(* Logix 5000 project; controller PLC_MCC1300_75F1 vendor 1 type 14 code 166 rev 32.11; software revision 32.04; part 50 of 83 *)
(* tags used below, declared in another part *)
   CM_ConveyorStackerToLine_JS1_Sync : CM_ConveyorStackerToLine;
   CONST_dDest_Cullet : DINT;
   CONST_dDest_Stk : DINT;
   CONST_rgdDestMask : DINT[32];   // Destination Mask
   Convoy_SL_DATA_NULL : UDT_Convoy_SL;
   GP_CheckIdPlatePresent : GP_CheckIdPlatePresent;
   GP_InvertCapxLite : GP_InvertCapxLite;
   GP_OB_InitializeMain : GP_OB_Initialize;
   GP_RampSpace : GP_RampSpace;
   Gp_SpaceConvUtilities_V1 : GP_SpaceConvUtilities_V1;
   M310B : MAC_Conveyor;
   M310B_ALM : MAC_Conveyor_ALM;
   M310B_Data : UDT_Convoy_SL;
   M310B_HMR : MAC_Conveyor_HMR;
   M310B_HMW : MAC_Conveyor_HMW;
   M310B_SpaceConv_Utilities : SpaceConv_Utilities;
   M310B_xPlateCullet : BOOL;
   M310Popup : MAC_Popup_ZC[2];
   M310Popup_SL_DATA : UDT_Convoy_SL;
   M311 : MAC_Conveyor;
   M311_Data : UDT_Convoy_SL;
   M311_SpaceConv_Utilities : SpaceConv_Utilities;
   M311_SpaceConvUtilities : SpaceConv_Utilities;
   M312 : MAC_Conveyor_Single;
   O : INT[128];
   TMP_d : DINT;
   TMP_dConveyorNumberForZoneCleaning : DINT;
   TMP_dDecelerationPositionEndConveyor : DINT;
   TMP_dHeadPosition : DINT;
   TMP_dOffsetLoadUnload_cmm : DINT;
   TMP_dPhEndPosition_cmm : DINT;
   TMP_dTailPosition : DINT;
   TMP_rgxId : DINT[10];
   TMP_SendToCullet : BOOL;
   TMP_xConveyorInvolvedInCleaning : BOOL;
   TMP_xConveyorOfStartCleaning : BOOL;
   TMP_xCulletPresent : BOOL;
   TMP_xEnableLoadUnload : BOOL;
   TMP_xEnableZoneCleaning : BOOL;
   TMP_xLiteThisDestPresent : BOOL;
   TMP_xReqUnpack : BOOL;
   xAlwaysOFF : BOOL;
   xAlwaysON : BOOL;
   Z401 : MAC_Zone;
   Z401_HMR : MAC_Zone_HMR;
   Z401_HMW : MAC_Zone_HMW;
(* MainProgram, continued *)

ROUTINE M310B_Logic   (* ladder *)
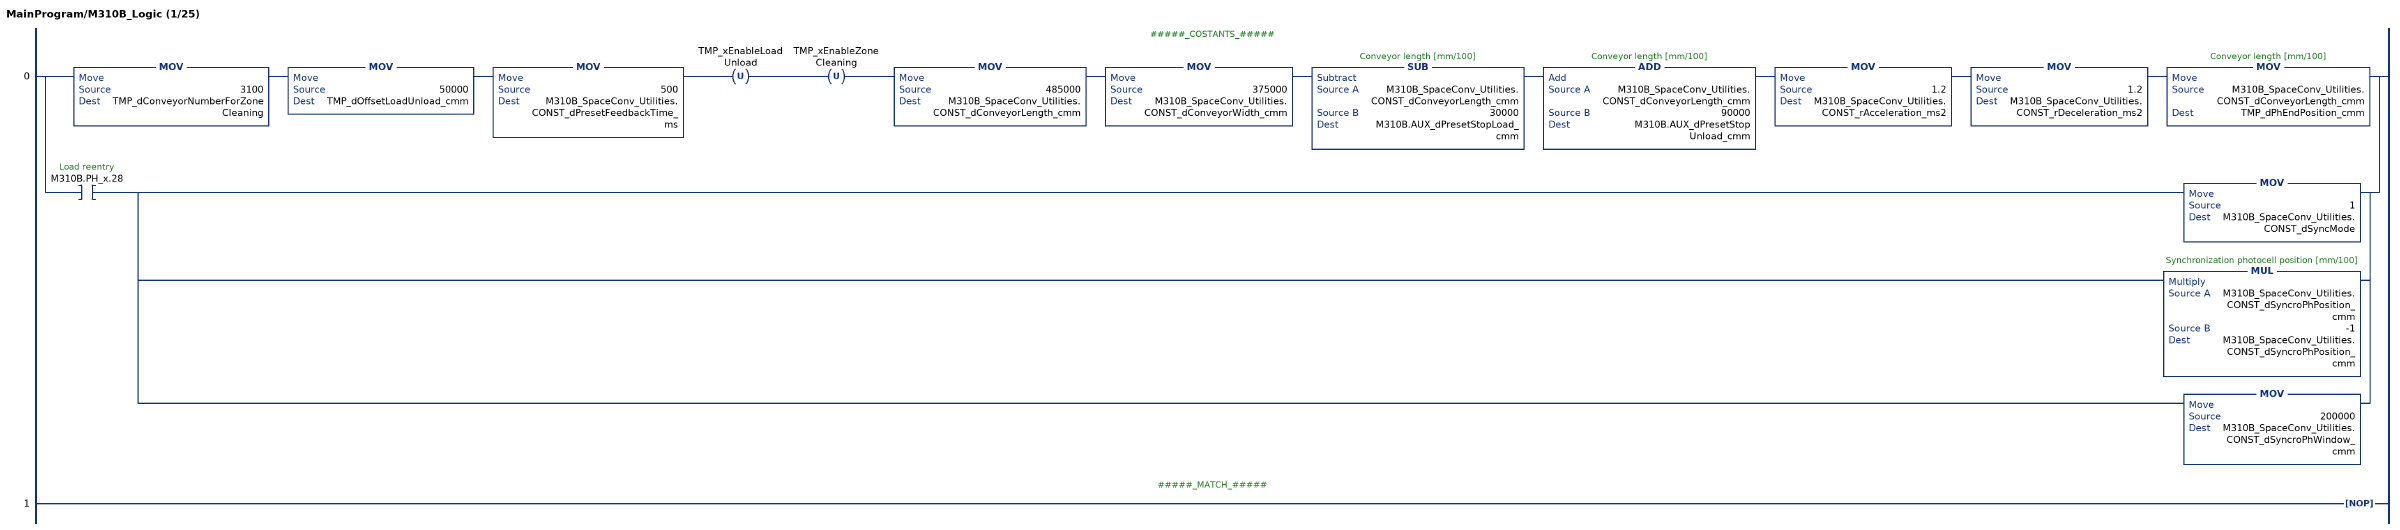
   // #####_COSTANTS_#####
   0: [MOV(3100,TMP_dConveyorNumberForZoneCleaning) MOV(50000,TMP_dOffsetLoadUnload_cmm) MOV(500,M310B_SpaceConv_Utilities.CONST_dPresetFeedbackTime_ms) OTU(TMP_xEnableLoadUnload) OTU(TMP_xEnableZoneCleaning) MOV(485000,M310B_SpaceConv_Utilities.CONST_dConveyorLength_cmm) MOV(375000,M310B_SpaceConv_Utilities.CONST_dConveyorWidth_cmm) SUB(M310B_SpaceConv_Utilities.CONST_dConveyorLength_cmm,30000,M310B.AUX_dPresetStopLoad_cmm) ADD(M310B_SpaceConv_Utilities.CONST_dConveyorLength_cmm,90000,M310B.AUX_dPresetStopUnload_cmm) MOV(1.2,M310B_SpaceConv_Utilities.CONST_rAcceleration_ms2) MOV(1.2,M310B_SpaceConv_Utilities.CONST_rDeceleration_ms2) MOV(M310B_SpaceConv_Utilities.CONST_dConveyorLength_cmm,TMP_dPhEndPosition_cmm) ,XIC(M310B.PH_x.28) [MOV(1,M310B_SpaceConv_Utilities.CONST_dSyncMode) ,MUL(M310B_SpaceConv_Utilities.CONST_dSyncroPhPosition_cmm,-1,M310B_SpaceConv_Utilities.CONST_dSyncroPhPosition_cmm) ,MOV(200000,M310B_SpaceConv_Utilities.CONST_dSyncroPhWindow_cmm) ] ];
   // #####_MATCH_#####
   1: NOP();
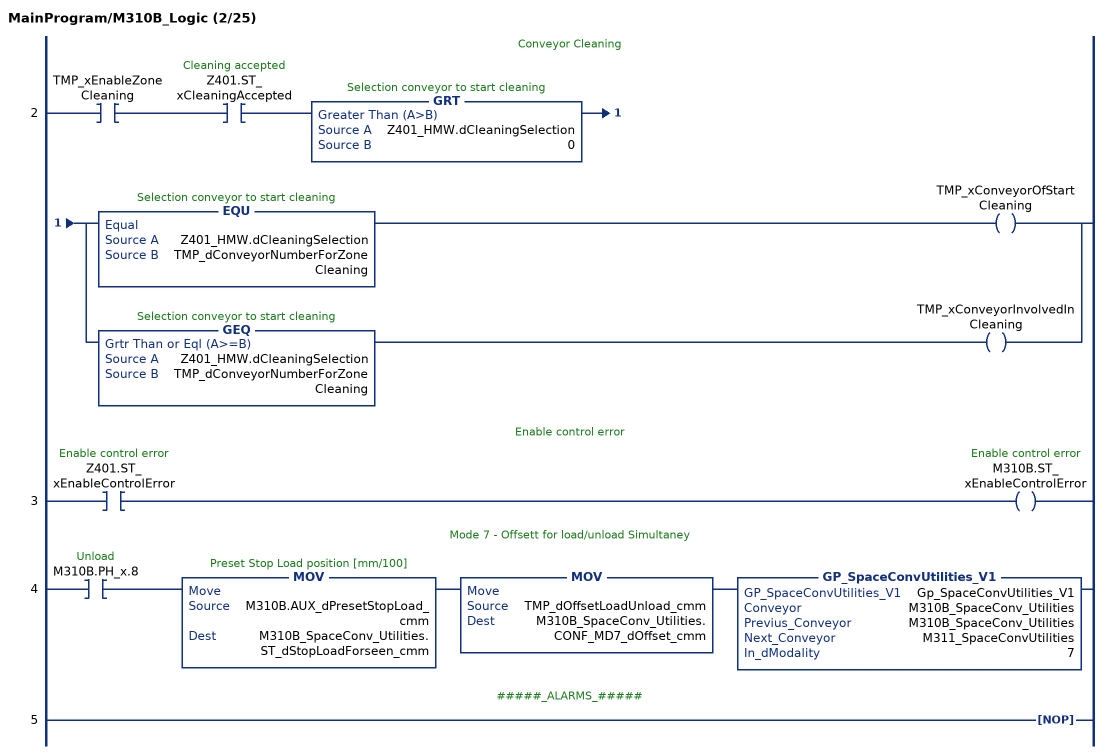
   // Conveyor Cleaning
   2: XIC(TMP_xEnableZoneCleaning)XIC(Z401.ST_xCleaningAccepted)GRT(Z401_HMW.dCleaningSelection,0)[EQU(Z401_HMW.dCleaningSelection,TMP_dConveyorNumberForZoneCleaning) OTE(TMP_xConveyorOfStartCleaning) ,GEQ(Z401_HMW.dCleaningSelection,TMP_dConveyorNumberForZoneCleaning) OTE(TMP_xConveyorInvolvedInCleaning) ];
   // Enable control error
   3: XIC(Z401.ST_xEnableControlError)OTE(M310B.ST_xEnableControlError);
   // Mode 7 - Offsett for load/unload Simultaney
   4: XIC(M310B.PH_x.8)MOV(M310B.AUX_dPresetStopLoad_cmm,M310B_SpaceConv_Utilities.ST_dStopLoadForseen_cmm)MOV(TMP_dOffsetLoadUnload_cmm,M310B_SpaceConv_Utilities.CONF_MD7_dOffset_cmm)GP_SpaceConvUtilities_V1(Gp_SpaceConvUtilities_V1,M310B_SpaceConv_Utilities,M310B_SpaceConv_Utilities,M311_SpaceConvUtilities,7);
   // #####_ALARMS_#####
   5: NOP();
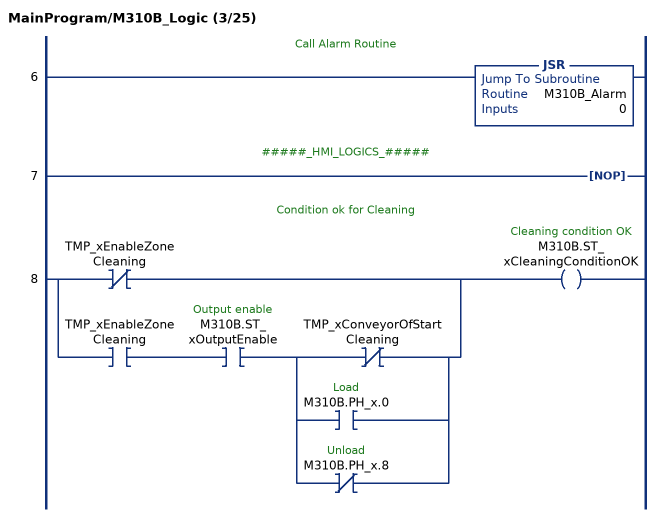
   // Call Alarm Routine
   6: JSR(M310B_Alarm,0);
   // #####_HMI_LOGICS_#####
   7: NOP();
   // Condition ok for Cleaning
   8: [XIO(TMP_xEnableZoneCleaning) ,XIC(TMP_xEnableZoneCleaning) XIC(M310B.ST_xOutputEnable) [XIO(TMP_xConveyorOfStartCleaning) ,XIC(M310B.PH_x.0) ,XIO(M310B.PH_x.8) ] ]OTE(M310B.ST_xCleaningConditionOK);
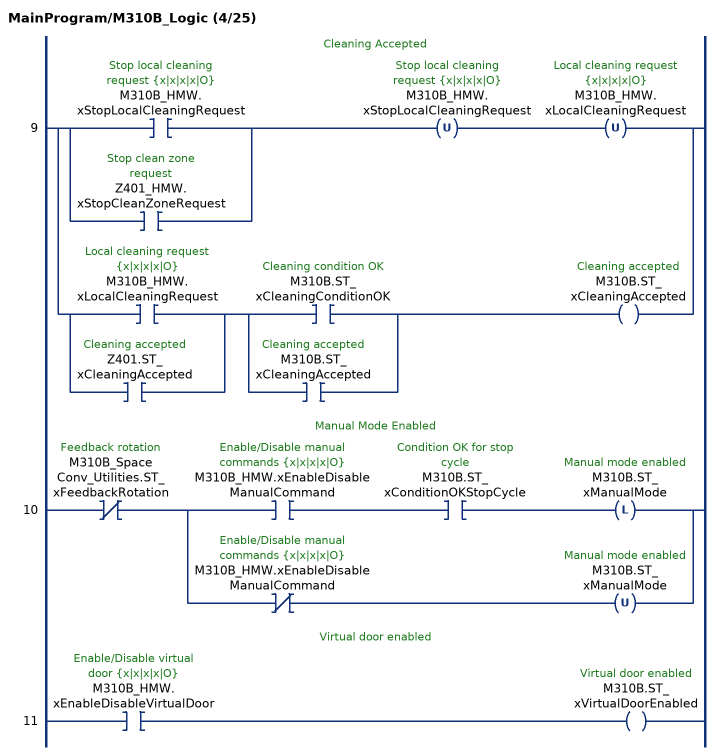
   // Cleaning Accepted
   9: [[XIC(M310B_HMW.xStopLocalCleaningRequest) ,XIC(Z401_HMW.xStopCleanZoneRequest) ] OTU(M310B_HMW.xStopLocalCleaningRequest) OTU(M310B_HMW.xLocalCleaningRequest) ,[XIC(M310B_HMW.xLocalCleaningRequest) ,XIC(Z401.ST_xCleaningAccepted) ] [XIC(M310B.ST_xCleaningConditionOK) ,XIC(M310B.ST_xCleaningAccepted) ] OTE(M310B.ST_xCleaningAccepted) ];
   // Manual Mode Enabled
   10: XIO(M310B_SpaceConv_Utilities.ST_xFeedbackRotation)[XIC(M310B_HMW.xEnableDisableManualCommand) XIC(M310B.ST_xConditionOKStopCycle) OTL(M310B.ST_xManualMode) ,XIO(M310B_HMW.xEnableDisableManualCommand) OTU(M310B.ST_xManualMode) ];
   // Virtual door enabled
   11: XIC(M310B_HMW.xEnableDisableVirtualDoor)OTE(M310B.ST_xVirtualDoorEnabled);
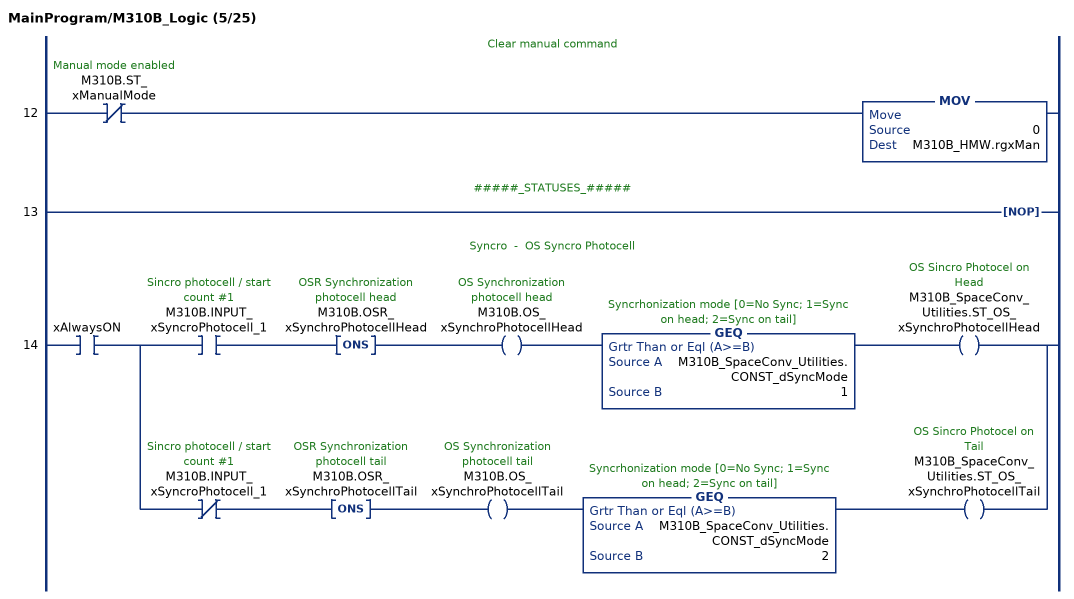
   // Clear manual command
   12: XIO(M310B.ST_xManualMode)MOV(0,M310B_HMW.rgxMan);
   // #####_STATUSES_#####
   13: NOP();
   // Syncro  -  OS Syncro Photocell
   14: XIC(xAlwaysON)[XIC(M310B.INPUT_xSyncroPhotocell_1) ONS(M310B.OSR_xSynchroPhotocellHead) OTE(M310B.OS_xSynchroPhotocellHead) GEQ(M310B_SpaceConv_Utilities.CONST_dSyncMode,1) OTE(M310B_SpaceConv_Utilities.ST_OS_xSynchroPhotocellHead) ,XIO(M310B.INPUT_xSyncroPhotocell_1) ONS(M310B.OSR_xSynchroPhotocellTail) OTE(M310B.OS_xSynchroPhotocellTail) GEQ(M310B_SpaceConv_Utilities.CONST_dSyncMode,2) OTE(M310B_SpaceConv_Utilities.ST_OS_xSynchroPhotocellTail) ];
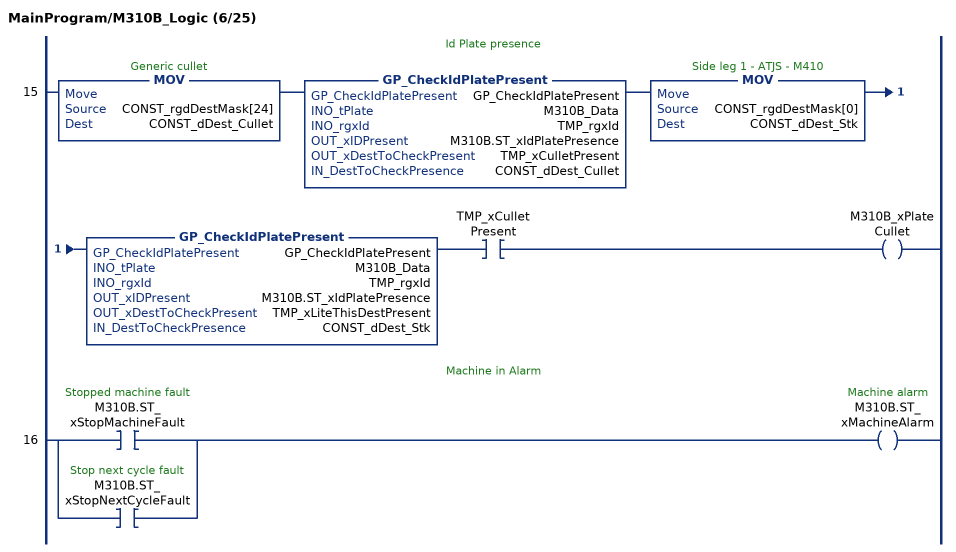
   // Id Plate presence
   15: MOV(CONST_rgdDestMask[24],CONST_dDest_Cullet)GP_CheckIdPlatePresent(GP_CheckIdPlatePresent,M310B_Data,TMP_rgxId,M310B.ST_xIdPlatePresence,TMP_xCulletPresent,CONST_dDest_Cullet)MOV(CONST_rgdDestMask[0],CONST_dDest_Stk)GP_CheckIdPlatePresent(GP_CheckIdPlatePresent,M310B_Data,TMP_rgxId,M310B.ST_xIdPlatePresence,TMP_xLiteThisDestPresent,CONST_dDest_Stk)XIC(TMP_xCulletPresent)OTE(M310B_xPlateCullet);
   // Machine in Alarm
   16: [XIC(M310B.ST_xStopMachineFault) ,XIC(M310B.ST_xStopNextCycleFault) ]OTE(M310B.ST_xMachineAlarm);
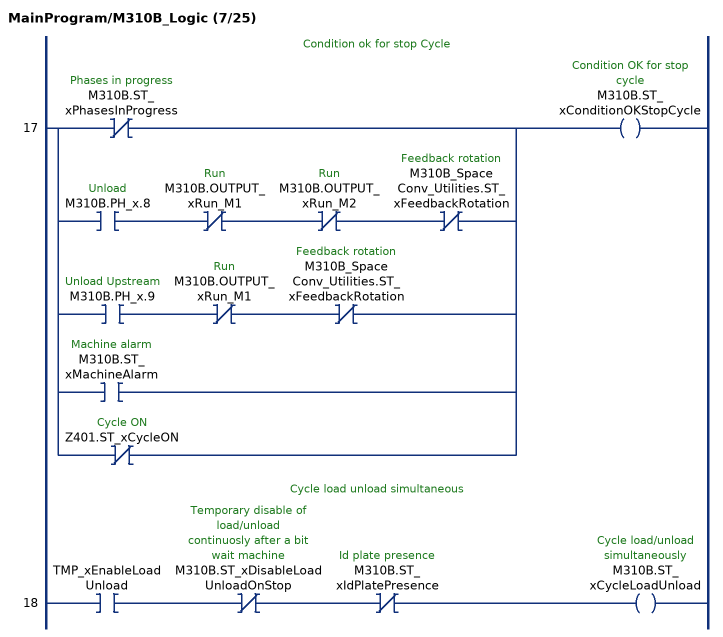
   // Condition ok for stop Cycle
   17: [XIO(M310B.ST_xPhasesInProgress) ,XIC(M310B.PH_x.8) XIO(M310B.OUTPUT_xRun_M1) XIO(M310B.OUTPUT_xRun_M2) XIO(M310B_SpaceConv_Utilities.ST_xFeedbackRotation) ,XIC(M310B.PH_x.9) XIO(M310B.OUTPUT_xRun_M1) XIO(M310B_SpaceConv_Utilities.ST_xFeedbackRotation) ,XIC(M310B.ST_xMachineAlarm) ,XIO(Z401.ST_xCycleON) ]OTE(M310B.ST_xConditionOKStopCycle);
   // Cycle load unload simultaneous
   18: XIC(TMP_xEnableLoadUnload)XIO(M310B.ST_xDisableLoadUnloadOnStop)XIO(M310B.ST_xIdPlatePresence)OTE(M310B.ST_xCycleLoadUnload);
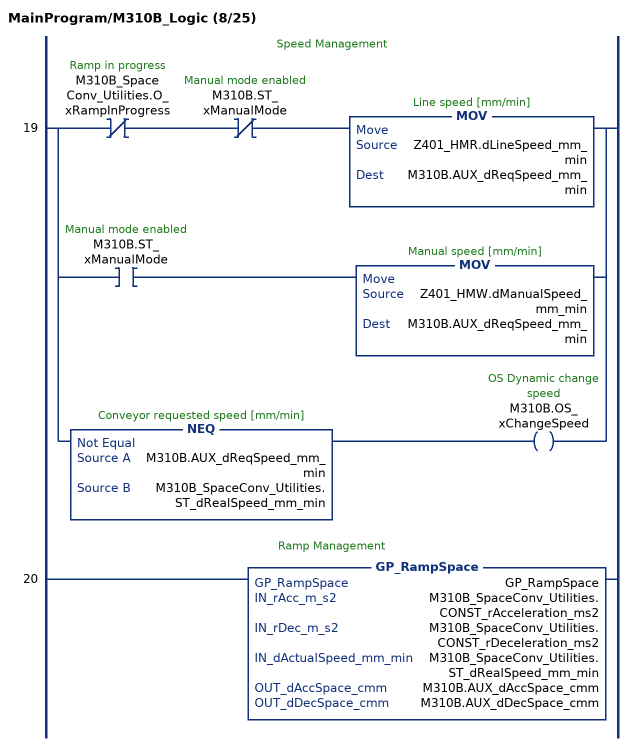
   // Speed Management
   19: [XIO(M310B_SpaceConv_Utilities.O_xRampInProgress) XIO(M310B.ST_xManualMode) MOV(Z401_HMR.dLineSpeed_mm_min,M310B.AUX_dReqSpeed_mm_min) ,XIC(M310B.ST_xManualMode) MOV(Z401_HMW.dManualSpeed_mm_min,M310B.AUX_dReqSpeed_mm_min) ,NEQ(M310B.AUX_dReqSpeed_mm_min,M310B_SpaceConv_Utilities.ST_dRealSpeed_mm_min) OTE(M310B.OS_xChangeSpeed) ];
   // Ramp Management
   20: GP_RampSpace(GP_RampSpace,M310B_SpaceConv_Utilities.CONST_rAcceleration_ms2,M310B_SpaceConv_Utilities.CONST_rDeceleration_ms2,M310B_SpaceConv_Utilities.ST_dRealSpeed_mm_min,M310B.AUX_dAccSpace_cmm,M310B.AUX_dDecSpace_cmm);
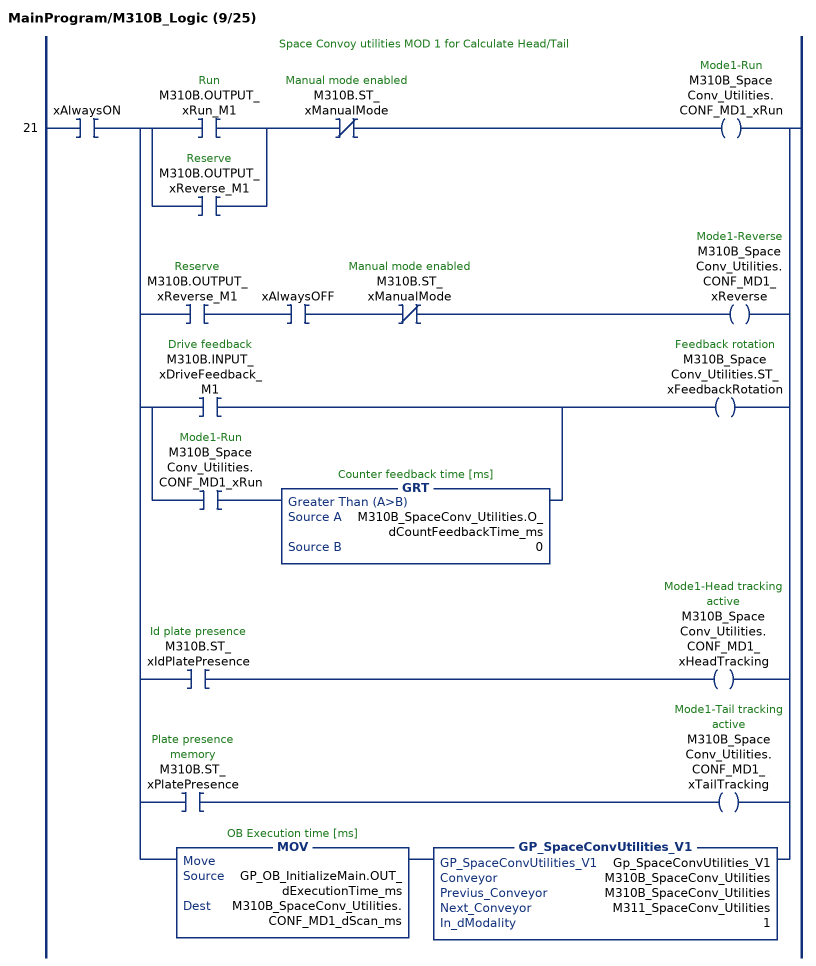
   // Space Convoy utilities MOD 1 for Calculate Head/Tail
   21: XIC(xAlwaysON)[[XIC(M310B.OUTPUT_xRun_M1) ,XIC(M310B.OUTPUT_xReverse_M1) ] XIO(M310B.ST_xManualMode) OTE(M310B_SpaceConv_Utilities.CONF_MD1_xRun) ,XIC(M310B.OUTPUT_xReverse_M1) XIC(xAlwaysOFF) XIO(M310B.ST_xManualMode) OTE(M310B_SpaceConv_Utilities.CONF_MD1_xReverse) ,[XIC(M310B.INPUT_xDriveFeedback_M1) ,XIC(M310B_SpaceConv_Utilities.CONF_MD1_xRun) GRT(M310B_SpaceConv_Utilities.O_dCountFeedbackTime_ms,0) ] OTE(M310B_SpaceConv_Utilities.ST_xFeedbackRotation) ,XIC(M310B.ST_xIdPlatePresence) OTE(M310B_SpaceConv_Utilities.CONF_MD1_xHeadTracking) ,XIC(M310B.ST_xPlatePresence) OTE(M310B_SpaceConv_Utilities.CONF_MD1_xTailTracking) ,MOV(GP_OB_InitializeMain.OUT_dExecutionTime_ms,M310B_SpaceConv_Utilities.CONF_MD1_dScan_ms) GP_SpaceConvUtilities_V1(Gp_SpaceConvUtilities_V1,M310B_SpaceConv_Utilities,M310B_SpaceConv_Utilities,M311_SpaceConv_Utilities,1) ];
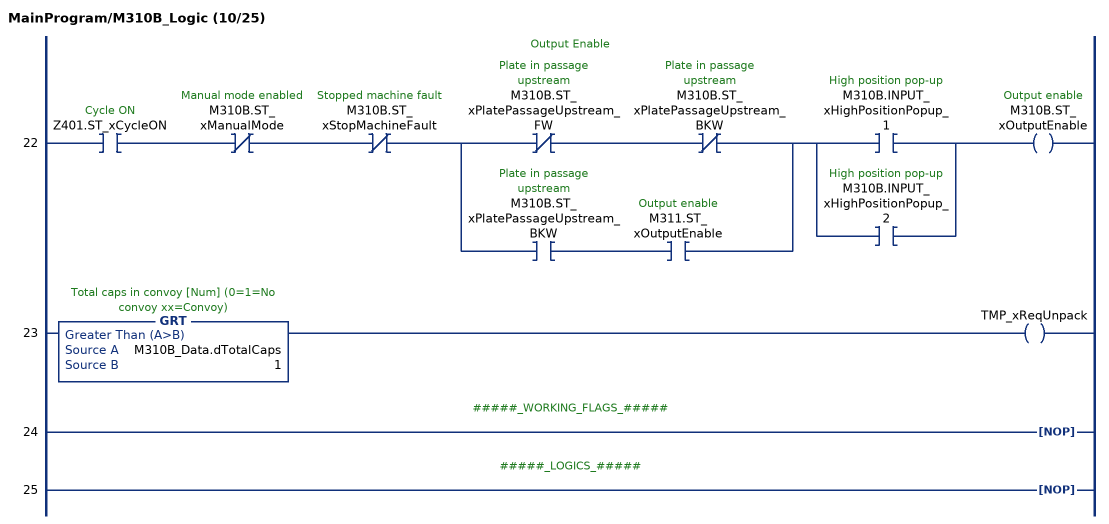
   // Output Enable
   22: XIC(Z401.ST_xCycleON)XIO(M310B.ST_xManualMode)XIO(M310B.ST_xStopMachineFault)[XIO(M310B.ST_xPlatePassageUpstream_FW) XIO(M310B.ST_xPlatePassageUpstream_BKW) ,XIC(M310B.ST_xPlatePassageUpstream_BKW) XIC(M311.ST_xOutputEnable) ][XIC(M310B.INPUT_xHighPositionPopup_1) ,XIC(M310B.INPUT_xHighPositionPopup_2) ]OTE(M310B.ST_xOutputEnable);
   23: GRT(M310B_Data.dTotalCaps,1)OTE(TMP_xReqUnpack);
   // #####_WORKING_FLAGS_#####
   24: NOP();
   // #####_LOGICS_#####
   25: NOP();
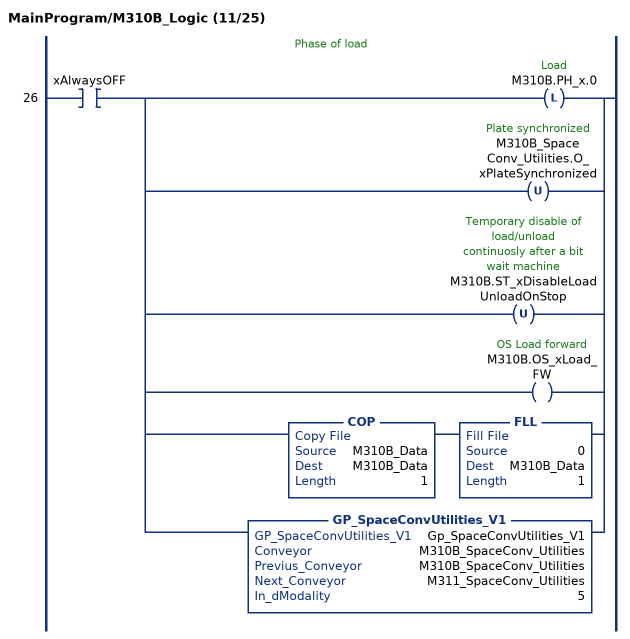
   // Phase of load
   26: XIC(xAlwaysOFF)[OTL(M310B.PH_x.0) ,OTU(M310B_SpaceConv_Utilities.O_xPlateSynchronized) ,OTU(M310B.ST_xDisableLoadUnloadOnStop) ,OTE(M310B.OS_xLoad_FW) ,COP(M310B_Data,M310B_Data,1) FLL(0,M310B_Data,1) ,GP_SpaceConvUtilities_V1(Gp_SpaceConvUtilities_V1,M310B_SpaceConv_Utilities,M310B_SpaceConv_Utilities,M311_SpaceConv_Utilities,5) ];
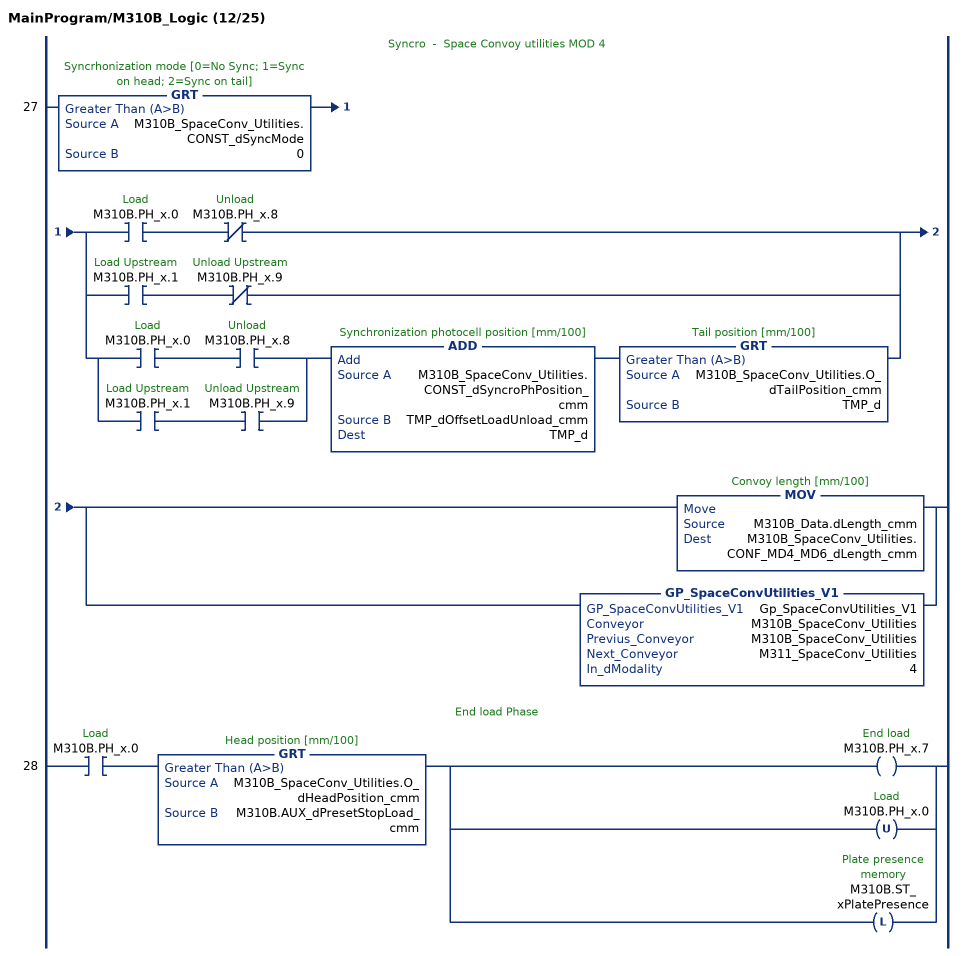
   // Syncro  -  Space Convoy utilities MOD 4
   27: GRT(M310B_SpaceConv_Utilities.CONST_dSyncMode,0)[[XIC(M310B.PH_x.0) XIO(M310B.PH_x.8) ,XIC(M310B.PH_x.1) XIO(M310B.PH_x.9) ] ,[XIC(M310B.PH_x.0) XIC(M310B.PH_x.8) ,XIC(M310B.PH_x.1) XIC(M310B.PH_x.9) ] ADD(M310B_SpaceConv_Utilities.CONST_dSyncroPhPosition_cmm,TMP_dOffsetLoadUnload_cmm,TMP_d) GRT(M310B_SpaceConv_Utilities.O_dTailPosition_cmm,TMP_d) ][MOV(M310B_Data.dLength_cmm,M310B_SpaceConv_Utilities.CONF_MD4_MD6_dLength_cmm) ,GP_SpaceConvUtilities_V1(Gp_SpaceConvUtilities_V1,M310B_SpaceConv_Utilities,M310B_SpaceConv_Utilities,M311_SpaceConv_Utilities,4) ];
   // End load Phase
   28: XIC(M310B.PH_x.0)GRT(M310B_SpaceConv_Utilities.O_dHeadPosition_cmm,M310B.AUX_dPresetStopLoad_cmm)[OTE(M310B.PH_x.7) ,OTU(M310B.PH_x.0) ,OTL(M310B.ST_xPlatePresence) ];